   	OWF_Key[32,16]:=227126216;
   	OWF_Key[33,13]:=74826149;
   	OWF_Key[33,14]:=1639015971;
   	OWF_Key[33,15]:=305196101;
   	OWF_Key[33,16]:=716882039;
   	OWF_Key[34,13]:=380880877;
   	OWF_Key[34,14]:=11839263;
   	OWF_Key[34,15]:=1373141717;
   	OWF_Key[34,16]:=532627490;
   	OWF_Key[35,13]:=93438529;
   	OWF_Key[35,14]:=35115978;
   	OWF_Key[35,15]:=1081533615;
   	OWF_Key[35,16]:=1111729827;
   	OWF_Key[36,13]:=380331581;
   	OWF_Key[36,14]:=1532456188;
   	OWF_Key[36,15]:=1939052724;
   	OWF_Key[36,16]:=1794611672;
   	OWF_Key[37,13]:=1819289397;
   	OWF_Key[37,14]:=1027002065;
   	OWF_Key[37,15]:=1244500467;
   	OWF_Key[37,16]:=936638688;
   	OWF_Key[38,13]:=1479190277;
   	OWF_Key[38,14]:=519596430;
   	OWF_Key[38,15]:=1911107362;
   	OWF_Key[38,16]:=435044551;
   	OWF_Key[39,13]:=917290529;
   	OWF_Key[39,14]:=1617052636;
   	OWF_Key[39,15]:=606522633;
   	OWF_Key[39,16]:=1781888676;
   	OWF_Key[40,13]:=1628193547;
   	OWF_Key[40,14]:=89927245;
   	OWF_Key[40,15]:=820592385;
   	OWF_Key[40,16]:=524162027;
   	OWF_Key[41,13]:=699504604;
   	OWF_Key[41,14]:=2016929121;
   	OWF_Key[41,15]:=1410565984;
   	OWF_Key[41,16]:=1344454938;
   	OWF_Key[42,13]:=346920590;
   	OWF_Key[42,14]:=546121623;
   	OWF_Key[42,15]:=1947269171;
   	OWF_Key[42,16]:=311947312;
   	OWF_Key[43,13]:=673700248;
   	OWF_Key[43,14]:=2041423853;
   	OWF_Key[43,15]:=875126022;
   	OWF_Key[43,16]:=1745165237;
   	OWF_Key[44,13]:=1753633549;
   	OWF_Key[44,14]:=1140321993;
   	OWF_Key[44,15]:=33633727;
   	OWF_Key[44,16]:=1343682688;
   	OWF_Key[45,13]:=299201156;
   	OWF_Key[45,14]:=293335340;
   	OWF_Key[45,15]:=666355512;
   	OWF_Key[45,16]:=1885349377;
   	OWF_Key[46,13]:=1439159427;
   	OWF_Key[46,14]:=628092582;
   	OWF_Key[46,15]:=1364839979;
   	OWF_Key[46,16]:=1866912;
   	OWF_Key[47,13]:=856720789;
   	OWF_Key[47,14]:=930916762;
   	OWF_Key[47,15]:=2123174806;
   	OWF_Key[47,16]:=1671058401;
   	OWF_Key[48,13]:=230854938;
   	OWF_Key[48,14]:=878476914;
   	OWF_Key[48,15]:=1158749479;
   	OWF_Key[48,16]:=1143227675;
   	OWF_Key[49,13]:=2073892953;
   	OWF_Key[49,14]:=1273666786;
   	OWF_Key[49,15]:=2144362013;
   	OWF_Key[49,16]:=1099736956;
   	OWF_Key[50,13]:=874888610;
   	OWF_Key[50,14]:=1873711650;
   	OWF_Key[50,15]:=1719753255;
   	OWF_Key[50,16]:=1680711035;
   	OWF_Key[51,13]:=1361816747;
   	OWF_Key[51,14]:=1994614458;
   	OWF_Key[51,15]:=1199333913;
   	OWF_Key[51,16]:=1830471925;
   	OWF_Key[52,13]:=1995713668;
   	OWF_Key[52,14]:=919849947;
   	OWF_Key[52,15]:=767203999;
   	OWF_Key[52,16]:=1950347560;
   	OWF_Key[53,13]:=1787066567;
   	OWF_Key[53,14]:=1641494518;
   	OWF_Key[53,15]:=2137169354;
   	OWF_Key[53,16]:=1052747155;
   	OWF_Key[54,13]:=2054621143;
   	OWF_Key[54,14]:=1974715107;
   	OWF_Key[54,15]:=2111338725;
   	OWF_Key[54,16]:=1642760447;
   	OWF_Key[55,13]:=315851187;
   	OWF_Key[55,14]:=1955885849;
   	OWF_Key[55,15]:=2037754524;
   	OWF_Key[55,16]:=1309783764;
   	OWF_Key[56,13]:=629952185;
   	OWF_Key[56,14]:=210914935;
   	OWF_Key[56,15]:=1623244036;
   	OWF_Key[56,16]:=1765475415;
   	OWF_Key[57,13]:=857435203;
   	OWF_Key[57,14]:=206048520;
   	OWF_Key[57,15]:=369910258;
   	OWF_Key[57,16]:=1843731464;
   	OWF_Key[58,13]:=324501666;
   	OWF_Key[58,14]:=1733381472;
   	OWF_Key[58,15]:=1847843539;
   	OWF_Key[58,16]:=1608870174;
   	OWF_Key[59,13]:=1465774380;
   	OWF_Key[59,14]:=1286619525;
   	OWF_Key[59,15]:=573519412;
   	OWF_Key[59,16]:=1150347743;
   	OWF_Key[60,13]:=2015895654;
   	OWF_Key[60,14]:=201882130;
   	OWF_Key[60,15]:=1496789631;
   	OWF_Key[60,16]:=753620274;
   	OWF_Key[61,13]:=258623275;
   	OWF_Key[61,14]:=542640591;
   	OWF_Key[61,15]:=1506681182;
   	OWF_Key[61,16]:=1854703257;
   	OWF_Key[62,13]:=1141501595;
   	OWF_Key[62,14]:=1968246431;
   	OWF_Key[62,15]:=1731135653;
   	OWF_Key[62,16]:=2019442968;
   	OWF_Key[63,13]:=1282787873;
   	OWF_Key[63,14]:=579188533;
   	OWF_Key[63,15]:=1379806521;
   	OWF_Key[63,16]:=1195986330;
   	OWF_Key[64,13]:=1760745701;
   	OWF_Key[64,14]:=796682114;
   	OWF_Key[64,15]:=503806046;
   	OWF_Key[64,16]:=1014065369;
   	OWF_Key[65,13]:=744789352;
   	OWF_Key[65,14]:=1669355124;
   	OWF_Key[65,15]:=1249003689;
   	OWF_Key[65,16]:=446383216;
   	OWF_Key[66,13]:=1359397698;
   	OWF_Key[66,14]:=157427355;
   	OWF_Key[66,15]:=488697501;
   	OWF_Key[66,16]:=1040142022;
   	OWF_Key[67,13]:=881757290;
   	OWF_Key[67,14]:=965262803;
   	OWF_Key[67,15]:=1915722473;
   	OWF_Key[67,16]:=656835267;
   	OWF_Key[68,13]:=933499237;
   	OWF_Key[68,14]:=1187531747;
   	OWF_Key[68,15]:=197012920;
   	OWF_Key[68,16]:=274156957;
   	OWF_Key[69,13]:=1435849115;
   	OWF_Key[69,14]:=207728093;
   	OWF_Key[69,15]:=1550339381;
   	OWF_Key[69,16]:=924520084;
   	OWF_Key[70,13]:=1792435968;
   	OWF_Key[70,14]:=290098793;
   	OWF_Key[70,15]:=823633063;
   	OWF_Key[70,16]:=905749060;
   	OWF_Key[71,13]:=1550939045;
   	OWF_Key[71,14]:=2047053549;
   	OWF_Key[71,15]:=613147771;
   	OWF_Key[71,16]:=1592945744;
   	OWF_Key[72,13]:=1671761274;
   	OWF_Key[72,14]:=1866470197;
   	OWF_Key[72,15]:=1595615064;
   	OWF_Key[72,16]:=1624872080;
   	OWF_Key[73,13]:=1330706500;
   	OWF_Key[73,14]:=995552984;
   	OWF_Key[73,15]:=1155990823;
   	OWF_Key[73,16]:=166888145;
   	OWF_Key[74,13]:=935434492;
   	OWF_Key[74,14]:=1004579779;
   	OWF_Key[74,15]:=441645409;
   	OWF_Key[74,16]:=1173860650;
   	OWF_Key[75,13]:=124465085;
   	OWF_Key[75,14]:=1848317617;
   	OWF_Key[75,15]:=774434070;
   	OWF_Key[75,16]:=1822370621;
   	OWF_Key[76,13]:=1955710974;
   	OWF_Key[76,14]:=963579763;
   	OWF_Key[76,15]:=1302080192;
   	OWF_Key[76,16]:=1915358529;
   	OWF_Key[77,13]:=510947175;
   	OWF_Key[77,14]:=1670479738;
   	OWF_Key[77,15]:=658812905;
   	OWF_Key[77,16]:=6552539;
   	OWF_Key[78,13]:=958044673;
   	OWF_Key[78,14]:=381647451;
   	OWF_Key[78,15]:=510842397;
   	OWF_Key[78,16]:=916863139;
   	OWF_Key[79,13]:=127497795;
   	OWF_Key[79,14]:=806273643;
   	OWF_Key[79,15]:=1652287201;
   	OWF_Key[79,16]:=1761646512;
   	OWF_Key[80,13]:=1319108753;
   	OWF_Key[80,14]:=119208384;
   	OWF_Key[80,15]:=1872549858;
   	OWF_Key[80,16]:=1745731921;
   	OWF_Key[81,13]:=1435598528;
   	OWF_Key[81,14]:=571194510;
   	OWF_Key[81,15]:=191567415;
   	OWF_Key[81,16]:=217112706;
   	OWF_Key[82,13]:=1754599579;
   	OWF_Key[82,14]:=514829758;
   	OWF_Key[82,15]:=242412916;
   	OWF_Key[82,16]:=1451035335;
   	OWF_Key[83,13]:=1055894451;
   	OWF_Key[83,14]:=153938916;
   	OWF_Key[83,15]:=1360024240;
   	OWF_Key[83,16]:=398108754;
   	OWF_Key[84,13]:=1483905120;
   	OWF_Key[84,14]:=117806243;
   	OWF_Key[84,15]:=822813432;
   	OWF_Key[84,16]:=422563876;
   	OWF_Key[85,13]:=162587349;
   	OWF_Key[85,14]:=478421491;
   	OWF_Key[85,15]:=1015415493;
   	OWF_Key[85,16]:=1830070223;
   	OWF_Key[86,13]:=334994722;
   	OWF_Key[86,14]:=1913921160;
   	OWF_Key[86,15]:=1114283805;
   	OWF_Key[86,16]:=1127178650;
   	OWF_Key[87,13]:=1107170890;
   	OWF_Key[87,14]:=2012352564;
   	OWF_Key[87,15]:=57491098;
   	OWF_Key[87,16]:=1031931037;
   	OWF_Key[88,13]:=1840152318;
   	OWF_Key[88,14]:=1439707080;
   	OWF_Key[88,15]:=1204125942;
   	OWF_Key[88,16]:=460202532;
   	OWF_Key[89,13]:=357664832;
   	OWF_Key[89,14]:=651670053;
   	OWF_Key[89,15]:=949523032;
   	OWF_Key[89,16]:=30336271;
   	OWF_Key[90,13]:=1537181786;
   	OWF_Key[90,14]:=385729653;
   	OWF_Key[90,15]:=702817811;
   	OWF_Key[90,16]:=506086235;
   	OWF_Key[91,13]:=140712957;
   	OWF_Key[91,14]:=1989169662;
   	OWF_Key[91,15]:=1948213053;
   	OWF_Key[91,16]:=1066195582;
   	OWF_Key[92,13]:=1080088464;
   	OWF_Key[92,14]:=463170373;
   	OWF_Key[92,15]:=323347074;
   	OWF_Key[92,16]:=1133893629;
   	OWF_Key[93,13]:=908912253;
   	OWF_Key[93,14]:=551968720;
   	OWF_Key[93,15]:=1980909314;
   	OWF_Key[93,16]:=1712465128;
   	OWF_Key[94,13]:=1085647434;
   	OWF_Key[94,14]:=1044237653;
   	OWF_Key[94,15]:=1675868506;
   	OWF_Key[94,16]:=323851357;
   	OWF_Key[95,13]:=898355252;
   	OWF_Key[95,14]:=1501587080;
   	OWF_Key[95,15]:=1296328976;
   	OWF_Key[95,16]:=858795092;
   	OWF_Key[96,13]:=1480170052;
   	OWF_Key[96,14]:=1561016974;
   	OWF_Key[96,15]:=388658317;
   	OWF_Key[96,16]:=1336155871;
   	OWF_Key[97,13]:=347985099;
   	OWF_Key[97,14]:=1819162848;
   	OWF_Key[97,15]:=1472264812;
   	OWF_Key[97,16]:=638122137;
   	OWF_Key[98,13]:=1693384262;
   	OWF_Key[98,14]:=287561249;
   	OWF_Key[98,15]:=248517399;
   	OWF_Key[98,16]:=2033544562;
   	OWF_Key[99,13]:=440390558;
   	OWF_Key[99,14]:=1349263930;
   	OWF_Key[99,15]:=1752934582;
   	OWF_Key[99,16]:=1828420687;
   	OWF_Key[100,13]:=1779162509;
   	OWF_Key[100,14]:=147277535;
   	OWF_Key[100,15]:=1591203745;
   	OWF_Key[100,16]:=1387986523;
   	OWF_Key[101,13]:=893571876;
   	OWF_Key[101,14]:=1470481068;
   	OWF_Key[101,15]:=539793699;
   	OWF_Key[101,16]:=37186580;
   	OWF_Key[102,13]:=1710752197;
   	OWF_Key[102,14]:=1484165743;
   	OWF_Key[102,15]:=502723645;
   	OWF_Key[102,16]:=1327015877;
   	OWF_Key[103,13]:=812458487;
   	OWF_Key[103,14]:=1628876014;
   	OWF_Key[103,15]:=1328316236;
   	OWF_Key[103,16]:=2054343353;
   	OWF_Key[104,13]:=1919425969;
   	OWF_Key[104,14]:=896029992;
   	OWF_Key[104,15]:=1110917444;
   	OWF_Key[104,16]:=425290322;
   	OWF_Key[105,13]:=1924264538;
   	OWF_Key[105,14]:=1216674049;
   	OWF_Key[105,15]:=1533302189;
   	OWF_Key[105,16]:=2115098790;
   	OWF_Key[106,13]:=444126867;
   	OWF_Key[106,14]:=1038812109;
   	OWF_Key[106,15]:=1620113783;
   	OWF_Key[106,16]:=1670203207;
   	OWF_Key[107,13]:=853022640;
   	OWF_Key[107,14]:=1446113967;
   	OWF_Key[107,15]:=331193698;
   	OWF_Key[107,16]:=36897127;
   	OWF_Key[108,13]:=1772607745;
   	OWF_Key[108,14]:=278613042;
   	OWF_Key[108,15]:=1641923280;
   	OWF_Key[108,16]:=901128481;
   	OWF_Key[109,13]:=462107376;
   	OWF_Key[109,14]:=1753942874;
   	OWF_Key[109,15]:=1420322543;
   	OWF_Key[109,16]:=1585835244;
   	OWF_Key[110,13]:=1025292899;
   	OWF_Key[110,14]:=377139452;
   	OWF_Key[110,15]:=960310545;
   	OWF_Key[110,16]:=1455759124;
   	OWF_Key[111,13]:=978224434;
   	OWF_Key[111,14]:=1769099284;
   	OWF_Key[111,15]:=1469343786;
   	OWF_Key[111,16]:=1894157702;
   	OWF_Key[112,13]:=1579369767;
   	OWF_Key[112,14]:=1221710590;
   	OWF_Key[112,15]:=27970548;
   	OWF_Key[112,16]:=475176021;
   	OWF_Key[113,13]:=1406741878;
   	OWF_Key[113,14]:=1391221516;
   	OWF_Key[113,15]:=973931164;
   	OWF_Key[113,16]:=935798566;
   	OWF_Key[114,13]:=1016826153;
   	OWF_Key[114,14]:=395417869;
   	OWF_Key[114,15]:=139427492;
   	OWF_Key[114,16]:=380613091;
   	OWF_Key[115,13]:=1199001387;
   	OWF_Key[115,14]:=1643051957;
   	OWF_Key[115,15]:=867375944;
   	OWF_Key[115,16]:=1768598715;
   	OWF_Key[116,13]:=1371985039;
   	OWF_Key[116,14]:=239918248;
   	OWF_Key[116,15]:=475467365;
   	OWF_Key[116,16]:=352629576;
   	OWF_Key[117,13]:=406649522;
   	OWF_Key[117,14]:=1022185637;
   	OWF_Key[117,15]:=924251933;
   	OWF_Key[117,16]:=58287288;
   	OWF_Key[118,13]:=1444359901;
   	OWF_Key[118,14]:=1004398136;
   	OWF_Key[118,15]:=305939276;
   	OWF_Key[118,16]:=13282582;
   	OWF_Key[119,13]:=1753624650;
   	OWF_Key[119,14]:=395513408;
   	OWF_Key[119,15]:=1423144984;
   	OWF_Key[119,16]:=1539743838;
   	OWF_Key[120,13]:=442395067;
   	OWF_Key[120,14]:=2018925503;
   	OWF_Key[120,15]:=953917663;
   	OWF_Key[120,16]:=1688609331;
   	OWF_Key[121,13]:=787971890;
   	OWF_Key[121,14]:=1620287384;
   	OWF_Key[121,15]:=256968225;
   	OWF_Key[121,16]:=1301956638;
   	OWF_Key[122,13]:=990668381;
   	OWF_Key[122,14]:=2018680738;
   	OWF_Key[122,15]:=915563951;
   	OWF_Key[122,16]:=1304501418;
   	OWF_Key[123,13]:=845352878;
   	OWF_Key[123,14]:=1326819379;
   	OWF_Key[123,15]:=973867524;
   	OWF_Key[123,16]:=1330778393;
   	OWF_Key[124,13]:=1212459966;
   	OWF_Key[124,14]:=331345962;
   	OWF_Key[124,15]:=1503496153;
   	OWF_Key[124,16]:=1881291653;
   	OWF_Key[125,13]:=275083085;
   	OWF_Key[125,14]:=1241962392;
   	OWF_Key[125,15]:=1663659714;
   	OWF_Key[125,16]:=359811177;
   	OWF_Key[126,13]:=469249223;
   	OWF_Key[126,14]:=862227537;
   	OWF_Key[126,15]:=1043658105;
   	OWF_Key[126,16]:=1730970707;
   	OWF_Key[127,13]:=1168087958;
   	OWF_Key[127,14]:=282353341;
   	OWF_Key[127,15]:=343861148;
   	OWF_Key[127,16]:=2052225671;
   	OWF_Key[128,13]:=1557870208;
   	OWF_Key[128,14]:=1209923749;
   	OWF_Key[128,15]:=1776967874;
   	OWF_Key[128,16]:=288485818;
   	OWF_Key[129,13]:=74300695;
   	OWF_Key[129,14]:=968535377;
   	OWF_Key[129,15]:=851571720;
   	OWF_Key[129,16]:=2094292864;
   	OWF_Key[130,13]:=102777636;
   	OWF_Key[130,14]:=410444836;
   	OWF_Key[130,15]:=1304169589;
   	OWF_Key[130,16]:=1061853872;
   	OWF_Key[131,13]:=935817478;
   	OWF_Key[131,14]:=1893612138;
   	OWF_Key[131,15]:=462395237;
   	OWF_Key[131,16]:=681940591;
   	OWF_Key[132,13]:=381652625;
   	OWF_Key[132,14]:=201502794;
   	OWF_Key[132,15]:=1754047887;
   	OWF_Key[132,16]:=311395707;
   	OWF_Key[133,13]:=346211181;
   	OWF_Key[133,14]:=2071318594;
   	OWF_Key[133,15]:=1513459740;
   	OWF_Key[133,16]:=1115232146;
   	OWF_Key[134,13]:=1598695163;
   	OWF_Key[134,14]:=1466344949;
   	OWF_Key[134,15]:=762229445;
   	OWF_Key[134,16]:=672484557;
   	OWF_Key[135,13]:=1650533870;
   	OWF_Key[135,14]:=746136511;
   	OWF_Key[135,15]:=1403884082;
   	OWF_Key[135,16]:=1128504661;
   	OWF_Key[136,13]:=1193152325;
   	OWF_Key[136,14]:=1642319657;
   	OWF_Key[136,15]:=764561960;
   	OWF_Key[136,16]:=1782348027;
   	OWF_Key[137,13]:=481612577;
   	OWF_Key[137,14]:=1117357605;
   	OWF_Key[137,15]:=1226367764;
   	OWF_Key[137,16]:=486415909;
   	OWF_Key[138,13]:=712276525;
   	OWF_Key[138,14]:=1231818236;
   	OWF_Key[138,15]:=889849699;
   	OWF_Key[138,16]:=1322456834;
   	OWF_Key[139,13]:=1658882780;
   	OWF_Key[139,14]:=299855880;
   	OWF_Key[139,15]:=457182275;
   	OWF_Key[139,16]:=375856677;
   	OWF_Key[140,13]:=1427201989;
   	OWF_Key[140,14]:=1842532478;
   	OWF_Key[140,15]:=2020223672;
   	OWF_Key[140,16]:=95163959;
   	OWF_Key[141,13]:=1076016553;
   	OWF_Key[141,14]:=1900141535;
   	OWF_Key[141,15]:=1257026434;
   	OWF_Key[141,16]:=909049460;
   	OWF_Key[142,13]:=372483116;
   	OWF_Key[142,14]:=152435569;
   	OWF_Key[142,15]:=1367585177;
   	OWF_Key[142,16]:=180714971;
   	OWF_Key[143,13]:=492180917;
   	OWF_Key[143,14]:=811497737;
   	OWF_Key[143,15]:=182411329;
   	OWF_Key[143,16]:=1448390505;
   	OWF_Key[144,13]:=1474316502;
   	OWF_Key[144,14]:=962265029;
   	OWF_Key[144,15]:=2143233034;
   	OWF_Key[144,16]:=86163621;
   	OWF_Key[145,13]:=22318259;
   	OWF_Key[145,14]:=464103670;
   	OWF_Key[145,15]:=9486028;
   	OWF_Key[145,16]:=165100234;
   	OWF_Key[146,13]:=1738036540;
   	OWF_Key[146,14]:=957495089;
   	OWF_Key[146,15]:=1871584640;
   	OWF_Key[146,16]:=88784541;
   	OWF_Key[147,13]:=326829794;
   	OWF_Key[147,14]:=1163466676;
   	OWF_Key[147,15]:=1555104822;
   	OWF_Key[147,16]:=2103407692;
   	OWF_Key[148,13]:=1529543674;
   	OWF_Key[148,14]:=71476052;
   	OWF_Key[148,15]:=1157626873;
   	OWF_Key[148,16]:=1806721818;
   	OWF_Key[149,13]:=1849787839;
   	OWF_Key[149,14]:=931886575;
   	OWF_Key[149,15]:=657127511;
   	OWF_Key[149,16]:=1271697867;
   	OWF_Key[150,13]:=1381878125;
   	OWF_Key[150,14]:=1019077359;
   	OWF_Key[150,15]:=1860188757;
   	OWF_Key[150,16]:=1322712000;
   	OWF_Key[151,13]:=648949296;
   	OWF_Key[151,14]:=99719;
   	OWF_Key[151,15]:=1175680819;
   	OWF_Key[151,16]:=1497980896;
   	OWF_Key[152,13]:=1625442764;
   	OWF_Key[152,14]:=277771665;
   	OWF_Key[152,15]:=939669588;
   	OWF_Key[152,16]:=1601021974;
   	OWF_Key[153,13]:=899912740;
   	OWF_Key[153,14]:=251847340;
   	OWF_Key[153,15]:=549386803;
   	OWF_Key[153,16]:=800804065;
   	OWF_Key[154,13]:=1113652973;
   	OWF_Key[154,14]:=47019578;
   	OWF_Key[154,15]:=1748787020;
   	OWF_Key[154,16]:=1741961176;
   	OWF_Key[155,13]:=16858922;
   	OWF_Key[155,14]:=993261889;
   	OWF_Key[155,15]:=391546459;
   	OWF_Key[155,16]:=1613990827;
   	OWF_Key[156,13]:=359980847;
   	OWF_Key[156,14]:=17310265;
   	OWF_Key[156,15]:=992777913;
   	OWF_Key[156,16]:=1166263769;
   	OWF_Key[157,13]:=1948582787;
   	OWF_Key[157,14]:=281935467;
   	OWF_Key[157,15]:=1445300746;
   	OWF_Key[157,16]:=1211611796;
   	OWF_Key[158,13]:=178475878;
   	OWF_Key[158,14]:=202525481;
   	OWF_Key[158,15]:=131006593;
   	OWF_Key[158,16]:=1956785807;
   	OWF_Key[159,13]:=1801698601;
   	OWF_Key[159,14]:=726011192;
   	OWF_Key[159,15]:=1429967167;
   	OWF_Key[159,16]:=120231144;
   	OWF_Key[160,13]:=1755934677;
   	OWF_Key[160,14]:=931127830;
   	OWF_Key[160,15]:=1573768517;
   	OWF_Key[160,16]:=194947820;
   	OWF_Key[161,13]:=340873654;
   	OWF_Key[161,14]:=859703477;
   	OWF_Key[161,15]:=714867666;
   	OWF_Key[161,16]:=1308970684;
   	OWF_Key[162,13]:=2033262093;
   	OWF_Key[162,14]:=135322483;
   	OWF_Key[162,15]:=181185071;
   	OWF_Key[162,16]:=1019448048;
   	OWF_Key[163,13]:=351815141;
   	OWF_Key[163,14]:=1349943554;
   	OWF_Key[163,15]:=1519426241;
   	OWF_Key[163,16]:=1730005141;
   	OWF_Key[164,13]:=895515385;
   	OWF_Key[164,14]:=759942475;
   	OWF_Key[164,15]:=1274974076;
   	OWF_Key[164,16]:=1778058459;
   	OWF_Key[165,13]:=1534002997;
   	OWF_Key[165,14]:=342683598;
   	OWF_Key[165,15]:=1325035008;
   	OWF_Key[165,16]:=541951738;
   	OWF_Key[166,13]:=1126159679;
   	OWF_Key[166,14]:=1135178360;
   	OWF_Key[166,15]:=171444871;
   	OWF_Key[166,16]:=1500118001;
   	OWF_Key[167,13]:=1319550750;
   	OWF_Key[167,14]:=1523155912;
   	OWF_Key[167,15]:=1894915506;
   	OWF_Key[167,16]:=46108147;
   	OWF_Key[168,13]:=891586055;
   	OWF_Key[168,14]:=1614220493;
   	OWF_Key[168,15]:=948985067;
   	OWF_Key[168,16]:=1008303949;
   	OWF_Key[169,13]:=714425471;
   	OWF_Key[169,14]:=404425965;
   	OWF_Key[169,15]:=1214720770;
   	OWF_Key[169,16]:=661094727;
   	OWF_Key[170,13]:=1417632945;
   	OWF_Key[170,14]:=1553623603;
   	OWF_Key[170,15]:=1142877093;
   	OWF_Key[170,16]:=1852102698;
   	OWF_Key[171,13]:=1325459671;
   	OWF_Key[171,14]:=1213428668;
   	OWF_Key[171,15]:=791381338;
   	OWF_Key[171,16]:=1093670539;
   	OWF_Key[172,13]:=67122307;
   	OWF_Key[172,14]:=722754093;
   	OWF_Key[172,15]:=1643848423;
   	OWF_Key[172,16]:=830718530;
   	OWF_Key[173,13]:=984850756;
   	OWF_Key[173,14]:=1149842119;
   	OWF_Key[173,15]:=171832428;
   	OWF_Key[173,16]:=2085848996;
   	OWF_Key[174,13]:=1995806419;
   	OWF_Key[174,14]:=811214497;
   	OWF_Key[174,15]:=1118289432;
   	OWF_Key[174,16]:=726787119;
   	OWF_Key[175,13]:=372222373;
   	OWF_Key[175,14]:=946921363;
   	OWF_Key[175,15]:=1763664559;
   	OWF_Key[175,16]:=1522951892;
   	OWF_Key[176,13]:=753425289;
   	OWF_Key[176,14]:=1971291402;
   	OWF_Key[176,15]:=1757383876;
   	OWF_Key[176,16]:=554600741;
   	OWF_Key[177,13]:=2116933958;
   	OWF_Key[177,14]:=684392856;
   	OWF_Key[177,15]:=1940251711;
   	OWF_Key[177,16]:=48359718;
   	OWF_Key[178,13]:=2028009177;
   	OWF_Key[178,14]:=48868902;
   	OWF_Key[178,15]:=89820102;
   	OWF_Key[178,16]:=1140097925;
   	OWF_Key[179,13]:=1985450806;
   	OWF_Key[179,14]:=1466515194;
   	OWF_Key[179,15]:=1981559753;
   	OWF_Key[179,16]:=465352035;
   	OWF_Key[180,13]:=1999606185;
   	OWF_Key[180,14]:=824765067;
   	OWF_Key[180,15]:=389379872;
   	OWF_Key[180,16]:=334105230;
   	OWF_Key[181,13]:=1123156879;
   	OWF_Key[181,14]:=1288903172;
   	OWF_Key[181,15]:=588243473;
   	OWF_Key[181,16]:=377190400;
   	OWF_Key[182,13]:=331455980;
   	OWF_Key[182,14]:=757004017;
   	OWF_Key[182,15]:=1679453652;
   	OWF_Key[182,16]:=953675030;
   	OWF_Key[183,13]:=319703761;
   	OWF_Key[183,14]:=686929024;
   	OWF_Key[183,15]:=1771394380;
   	OWF_Key[183,16]:=1146391459;
   	OWF_Key[184,13]:=64113331;
   	OWF_Key[184,14]:=1843233077;
   	OWF_Key[184,15]:=1054710883;
   	OWF_Key[184,16]:=16307061;
   	OWF_Key[185,13]:=577790918;
   	OWF_Key[185,14]:=769951951;
   	OWF_Key[185,15]:=36875238;
   	OWF_Key[185,16]:=969551747;
   	OWF_Key[186,13]:=1949099229;
   	OWF_Key[186,14]:=16345749;
   	OWF_Key[186,15]:=1812777874;
   	OWF_Key[186,16]:=1770825016;
   	OWF_Key[187,13]:=360969632;
   	OWF_Key[187,14]:=1677985071;
   	OWF_Key[187,15]:=1100521128;
   	OWF_Key[187,16]:=1658272940;
   	OWF_Key[188,13]:=1778139981;
   	OWF_Key[188,14]:=1202793776;
   	OWF_Key[188,15]:=17874512;
   	OWF_Key[188,16]:=2077025197;
   	OWF_Key[189,13]:=1605074632;
   	OWF_Key[189,14]:=735118058;
   	OWF_Key[189,15]:=2120994248;
   	OWF_Key[189,16]:=1327201891;
   	OWF_Key[190,13]:=2070065568;
   	OWF_Key[190,14]:=1393044672;
   	OWF_Key[190,15]:=976654796;
   	OWF_Key[190,16]:=1710671530;
   	OWF_Key[191,13]:=38568234;
   	OWF_Key[191,14]:=451698160;
   	OWF_Key[191,15]:=1261954091;
   	OWF_Key[191,16]:=249271037;
   	OWF_Key[192,13]:=1638949335;
   	OWF_Key[192,14]:=8243760;
   	OWF_Key[192,15]:=241234447;
   	OWF_Key[192,16]:=1227077516;
   	OWF_Key[193,13]:=989587635;
   	OWF_Key[193,14]:=1819989847;
   	OWF_Key[193,15]:=1332579048;
   	OWF_Key[193,16]:=53755968;
   	OWF_Key[194,13]:=100673663;
   	OWF_Key[194,14]:=1469329794;
   	OWF_Key[194,15]:=1436971146;
   	OWF_Key[194,16]:=929174323;
   	OWF_Key[195,13]:=577996306;
   	OWF_Key[195,14]:=1745684579;
   	OWF_Key[195,15]:=1996965839;
   	OWF_Key[195,16]:=1403732815;
   	OWF_Key[196,13]:=814419608;
   	OWF_Key[196,14]:=2103643129;
   	OWF_Key[196,15]:=335105042;
   	OWF_Key[196,16]:=565961710;
   	OWF_Key[197,13]:=202009593;
   	OWF_Key[197,14]:=930351125;
   	OWF_Key[197,15]:=1526609745;
   	OWF_Key[197,16]:=235969148;
   	OWF_Key[198,13]:=1626921131;
   	OWF_Key[198,14]:=161315506;
   	OWF_Key[198,15]:=767020089;
   	OWF_Key[198,16]:=624440912;
   	OWF_Key[199,13]:=684936633;
   	OWF_Key[199,14]:=1742723201;
   	OWF_Key[199,15]:=515114070;
   	OWF_Key[199,16]:=162561603;
   	OWF_Key[200,13]:=1845652691;
   	OWF_Key[200,14]:=1950369016;
   	OWF_Key[200,15]:=571396495;
   	OWF_Key[200,16]:=1488194196;
   	OWF_Key[201,13]:=1043958765;
   	OWF_Key[201,14]:=1442574514;
   	OWF_Key[201,15]:=298914684;
   	OWF_Key[201,16]:=486285287;
   	OWF_Key[202,13]:=1582775329;
   	OWF_Key[202,14]:=838793472;
   	OWF_Key[202,15]:=418382333;
   	OWF_Key[202,16]:=10776897;
   	OWF_Key[203,13]:=356986201;
   	OWF_Key[203,14]:=1108865874;
   	OWF_Key[203,15]:=1219664864;
   	OWF_Key[203,16]:=333594191;
   	OWF_Key[204,13]:=1541947490;
   	OWF_Key[204,14]:=1287551736;
   	OWF_Key[204,15]:=2059108066;
   	OWF_Key[204,16]:=1345707128;
   	OWF_Key[205,13]:=471367747;
   	OWF_Key[205,14]:=1525775149;
   	OWF_Key[205,15]:=1316108369;
   	OWF_Key[205,16]:=204019700;
   	OWF_Key[206,13]:=1473740948;
   	OWF_Key[206,14]:=286079449;
   	OWF_Key[206,15]:=1267750516;
   	OWF_Key[206,16]:=1937545157;
   	OWF_Key[207,13]:=2126324793;
   	OWF_Key[207,14]:=1789210342;
   	OWF_Key[207,15]:=501529746;
   	OWF_Key[207,16]:=2059785685;
   	OWF_Key[208,13]:=1274331883;
   	OWF_Key[208,14]:=968436149;
   	OWF_Key[208,15]:=1212562234;
   	OWF_Key[208,16]:=1455603155;
   	OWF_Key[209,13]:=92139053;
   	OWF_Key[209,14]:=992103779;
   	OWF_Key[209,15]:=1748163220;
   	OWF_Key[209,16]:=1233220835;
   	OWF_Key[210,13]:=259332684;
   	OWF_Key[210,14]:=2097850167;
   	OWF_Key[210,15]:=1049341383;
   	OWF_Key[210,16]:=714331988;
   	OWF_Key[211,13]:=1943218259;
   	OWF_Key[211,14]:=783610855;
   	OWF_Key[211,15]:=1161953504;
   	OWF_Key[211,16]:=1696436050;
   	OWF_Key[212,13]:=153726579;
   	OWF_Key[212,14]:=1993949032;
   	OWF_Key[212,15]:=281746886;
   	OWF_Key[212,16]:=2143629952;
   	OWF_Key[213,13]:=605671393;
   	OWF_Key[213,14]:=1472561361;
   	OWF_Key[213,15]:=1039695812;
   	OWF_Key[213,16]:=1849168053;
   	OWF_Key[214,13]:=1769778486;
   	OWF_Key[214,14]:=45741824;
   	OWF_Key[214,15]:=87024642;
   	OWF_Key[214,16]:=327652964;
   	OWF_Key[215,13]:=1490125572;
   	OWF_Key[215,14]:=1994649884;
   	OWF_Key[215,15]:=1234571844;
   	OWF_Key[215,16]:=920030323;
   	OWF_Key[216,13]:=2133174690;
   	OWF_Key[216,14]:=95558060;
   	OWF_Key[216,15]:=615326818;
   	OWF_Key[216,16]:=761728021;
   	OWF_Key[217,13]:=382282573;
   	OWF_Key[217,14]:=2017861784;
   	OWF_Key[217,15]:=1878700514;
   	OWF_Key[217,16]:=1515922417;
   	OWF_Key[218,13]:=1408298373;
   	OWF_Key[218,14]:=2039732974;
   	OWF_Key[218,15]:=1146678000;
   	OWF_Key[218,16]:=527275423;
   	OWF_Key[219,13]:=9291349;
   	OWF_Key[219,14]:=1702428079;
   	OWF_Key[219,15]:=340543343;
   	OWF_Key[219,16]:=1326649665;
   	OWF_Key[220,13]:=688341233;
   	OWF_Key[220,14]:=641189597;
   	OWF_Key[220,15]:=909299166;
   	OWF_Key[220,16]:=1752870415;
   	OWF_Key[221,13]:=1293014471;
   	OWF_Key[221,14]:=1168109613;
   	OWF_Key[221,15]:=1639198412;
   	OWF_Key[221,16]:=1211155230;
   	OWF_Key[222,13]:=1094302685;
   	OWF_Key[222,14]:=1748380807;
   	OWF_Key[222,15]:=740974356;
   	OWF_Key[222,16]:=981054882;
   	OWF_Key[223,13]:=1672948985;
   	OWF_Key[223,14]:=653486474;
   	OWF_Key[223,15]:=252491540;
   	OWF_Key[223,16]:=233857892;
   	OWF_Key[224,13]:=1488948359;
   	OWF_Key[224,14]:=855793400;
   	OWF_Key[224,15]:=299892487;
   	OWF_Key[224,16]:=955554724;
   	OWF_Key[225,13]:=1321934707;
   	OWF_Key[225,14]:=515714607;
   	OWF_Key[225,15]:=1346403512;
   	OWF_Key[225,16]:=540889864;
   	OWF_Key[226,13]:=760856919;
   	OWF_Key[226,14]:=452777885;
   	OWF_Key[226,15]:=152820366;
   	OWF_Key[226,16]:=158283786;
   	OWF_Key[227,13]:=1089442553;
   	OWF_Key[227,14]:=2136824552;
   	OWF_Key[227,15]:=492274941;
   	OWF_Key[227,16]:=1279116002;
   	OWF_Key[228,13]:=1639087779;
   	OWF_Key[228,14]:=1218708088;
   	OWF_Key[228,15]:=1350789742;
   	OWF_Key[228,16]:=266569552;
   	OWF_Key[229,13]:=63735330;
   	OWF_Key[229,14]:=1886757000;
   	OWF_Key[229,15]:=1923484766;
   	OWF_Key[229,16]:=1872440511;
   	OWF_Key[230,13]:=1943052252;
   	OWF_Key[230,14]:=1939759099;
   	OWF_Key[230,15]:=1108124166;
   	OWF_Key[230,16]:=1825389873;
   	OWF_Key[231,13]:=106697806;
   	OWF_Key[231,14]:=934330632;
   	OWF_Key[231,15]:=1226706106;
   	OWF_Key[231,16]:=1350717017;
   	OWF_Key[232,13]:=894995339;
   	OWF_Key[232,14]:=351973824;
   	OWF_Key[232,15]:=1915615287;
   	OWF_Key[232,16]:=1129455312;
   	OWF_Key[233,13]:=1606628665;
   	OWF_Key[233,14]:=792183115;
   	OWF_Key[233,15]:=655199967;
   	OWF_Key[233,16]:=466042394;
   	OWF_Key[234,13]:=265845209;
   	OWF_Key[234,14]:=1445558412;
   	OWF_Key[234,15]:=929515350;
   	OWF_Key[234,16]:=1736036285;
   	OWF_Key[235,13]:=1417713492;
   	OWF_Key[235,14]:=1710605342;
   	OWF_Key[235,15]:=153446933;
   	OWF_Key[235,16]:=200651284;
   	OWF_Key[236,13]:=1199064634;
   	OWF_Key[236,14]:=1304667317;
   	OWF_Key[236,15]:=1611340556;
   	OWF_Key[236,16]:=1688220347;
   	OWF_Key[237,13]:=1064686683;
   	OWF_Key[237,14]:=808058326;
   	OWF_Key[237,15]:=602176291;
   	OWF_Key[237,16]:=1592512372;
   	OWF_Key[238,13]:=188870782;
   	OWF_Key[238,14]:=699286542;
   	OWF_Key[238,15]:=740512834;
   	OWF_Key[238,16]:=805888291;
   	OWF_Key[239,13]:=2112249627;
   	OWF_Key[239,14]:=104687811;
   	OWF_Key[239,15]:=327040909;
   	OWF_Key[239,16]:=106310827;
   	OWF_Key[240,13]:=1922545948;
   	OWF_Key[240,14]:=1158736547;
   	OWF_Key[240,15]:=1646338950;
   	OWF_Key[240,16]:=302904535;
   	OWF_Key[241,13]:=1445166756;
   	OWF_Key[241,14]:=619904940;
   	OWF_Key[241,15]:=805963919;
   	OWF_Key[241,16]:=1775549581;
   	OWF_Key[242,13]:=461521008;
   	OWF_Key[242,14]:=1556197099;
   	OWF_Key[242,15]:=1292972172;
   	OWF_Key[242,16]:=1092790932;
   	OWF_Key[243,13]:=1366207430;
   	OWF_Key[243,14]:=1785310964;
   	OWF_Key[243,15]:=568468368;
   	OWF_Key[243,16]:=1252968121;
   	OWF_Key[244,13]:=973501638;
   	OWF_Key[244,14]:=859732749;
   	OWF_Key[244,15]:=1833062061;
   	OWF_Key[244,16]:=572987018;
   	OWF_Key[245,13]:=791865080;
   	OWF_Key[245,14]:=1765055225;
   	OWF_Key[245,15]:=310873594;
   	OWF_Key[245,16]:=589255605;
   	OWF_Key[246,13]:=1759833367;
   	OWF_Key[246,14]:=1618489300;
   	OWF_Key[246,15]:=830573894;
   	OWF_Key[246,16]:=1046861291;
   	OWF_Key[247,13]:=273538380;
   	OWF_Key[247,14]:=45619103;
   	OWF_Key[247,15]:=1158253128;
   	OWF_Key[247,16]:=142007761;
   	OWF_Key[248,13]:=307057508;
   	OWF_Key[248,14]:=1407424654;
   	OWF_Key[248,15]:=1570069593;
   	OWF_Key[248,16]:=832481957;
   	OWF_Key[249,13]:=962494443;
   	OWF_Key[249,14]:=1117874804;
   	OWF_Key[249,15]:=1823842561;
   	OWF_Key[249,16]:=1850442054;
   	OWF_Key[250,13]:=1442058163;
   	OWF_Key[250,14]:=1232560055;
   	OWF_Key[250,15]:=151821927;
   	OWF_Key[250,16]:=1056371398;
   	OWF_Key[251,13]:=332739772;
   	OWF_Key[251,14]:=2051033636;
   	OWF_Key[251,15]:=849642509;
   	OWF_Key[251,16]:=1992496557;
   	OWF_Key[252,13]:=1955024293;
   	OWF_Key[252,14]:=864654120;
   	OWF_Key[252,15]:=400202456;
   	OWF_Key[252,16]:=1469872697;
   	OWF_Key[253,13]:=1814679055;
   	OWF_Key[253,14]:=1018947711;
   	OWF_Key[253,15]:=414056628;
   	OWF_Key[253,16]:=1916175716;
   	OWF_Key[254,13]:=34988910;
   	OWF_Key[254,14]:=1068930085;
   	OWF_Key[254,15]:=1069419481;
   	OWF_Key[254,16]:=1329460403;
   	OWF_Key[255,13]:=629578987;
   	OWF_Key[255,14]:=1913112785;
   	OWF_Key[255,15]:=1118884227;
   	OWF_Key[255,16]:=660504630;
   	OWF_Key[256,13]:=1745889977;
   	OWF_Key[256,14]:=1744367642;
   	OWF_Key[256,15]:=1635265674;
   	OWF_Key[256,16]:=250591589;
   	OWF_Key[257,13]:=1359647390;
   	OWF_Key[257,14]:=335557629;
   	OWF_Key[257,15]:=272575744;
   	OWF_Key[257,16]:=782479111;
   	OWF_Key[258,13]:=1684017798;
   	OWF_Key[258,14]:=1849154465;
   	OWF_Key[258,15]:=131467400;
   	OWF_Key[258,16]:=244488627;
   	OWF_Key[259,13]:=41240583;
   	OWF_Key[259,14]:=963084835;
   	OWF_Key[259,15]:=844053562;
   	OWF_Key[259,16]:=1313394598;
   	OWF_Key[260,13]:=646795143;
   	OWF_Key[260,14]:=1614027852;
   	OWF_Key[260,15]:=2028202305;
   	OWF_Key[260,16]:=1145473513;
   	OWF_Key[261,13]:=16520506;
   	OWF_Key[261,14]:=1480547316;
   	OWF_Key[261,15]:=1576651890;
   	OWF_Key[261,16]:=326846098;
   	OWF_Key[262,13]:=274761447;
   	OWF_Key[262,14]:=981162513;
   	OWF_Key[262,15]:=960880365;
   	OWF_Key[262,16]:=535655077;
   	OWF_Key[263,13]:=815853165;
   	OWF_Key[263,14]:=965917766;
   	OWF_Key[263,15]:=1914171172;
   	OWF_Key[263,16]:=192053027;
   	OWF_Key[264,13]:=908824118;
   	OWF_Key[264,14]:=2075268001;
   	OWF_Key[264,15]:=314233580;
   	OWF_Key[264,16]:=1793819686;
   	OWF_Key[265,13]:=928633642;
   	OWF_Key[265,14]:=1394677407;
   	OWF_Key[265,15]:=381077257;
   	OWF_Key[265,16]:=1427933170;
   	OWF_Key[266,13]:=1325823149;
   	OWF_Key[266,14]:=326658029;
   	OWF_Key[266,15]:=1415638516;
   	OWF_Key[266,16]:=1370549208;
   	OWF_Key[267,13]:=91918653;
   	OWF_Key[267,14]:=1189442786;
   	OWF_Key[267,15]:=1488204864;
   	OWF_Key[267,16]:=739198522;
   	OWF_Key[268,13]:=1461502145;
   	OWF_Key[268,14]:=84921185;
   	OWF_Key[268,15]:=440014277;
   	OWF_Key[268,16]:=2099928856;
   	OWF_Key[269,13]:=1927983756;
   	OWF_Key[269,14]:=1119840967;
   	OWF_Key[269,15]:=388770855;
   	OWF_Key[269,16]:=1179250891;
   	OWF_Key[270,13]:=126605253;
   	OWF_Key[270,14]:=777231285;
   	OWF_Key[270,15]:=2005758675;
   	OWF_Key[270,16]:=1335960631;
   	OWF_Key[271,13]:=1845648579;
   	OWF_Key[271,14]:=380266852;
   	OWF_Key[271,15]:=248475413;
   	OWF_Key[271,16]:=331001610;
   	OWF_Key[272,13]:=605803683;
   	OWF_Key[272,14]:=607759287;
   	OWF_Key[272,15]:=665317173;
   	OWF_Key[272,16]:=1066666071;
   	OWF_Key[273,13]:=1398348673;
   	OWF_Key[273,14]:=848648801;
   	OWF_Key[273,15]:=867913242;
   	OWF_Key[273,16]:=138992559;
   	OWF_Key[274,13]:=610350804;
   	OWF_Key[274,14]:=523330815;
   	OWF_Key[274,15]:=1415166854;
   	OWF_Key[274,16]:=1770062347;
   	OWF_Key[275,13]:=835727048;
   	OWF_Key[275,14]:=35430845;
   	OWF_Key[275,15]:=596122974;
   	OWF_Key[275,16]:=684344241;
   	OWF_Key[276,13]:=78641305;
   	OWF_Key[276,14]:=788905719;
   	OWF_Key[276,15]:=880092642;
   	OWF_Key[276,16]:=1020585456;
   	OWF_Key[277,13]:=1110913439;
   	OWF_Key[277,14]:=1364792795;
   	OWF_Key[277,15]:=1384151855;
   	OWF_Key[277,16]:=1781215518;
   	OWF_Key[278,13]:=1664996503;
   	OWF_Key[278,14]:=1954790028;
   	OWF_Key[278,15]:=320064116;
   	OWF_Key[278,16]:=318277611;
   	OWF_Key[279,13]:=1474869755;
   	OWF_Key[279,14]:=1993904309;
   	OWF_Key[279,15]:=749636549;
   	OWF_Key[279,16]:=2065511657;
   	OWF_Key[280,13]:=903827560;
   	OWF_Key[280,14]:=1827376749;
   	OWF_Key[280,15]:=103307236;
   	OWF_Key[280,16]:=510364959;
   	OWF_Key[281,13]:=1734942199;
   	OWF_Key[281,14]:=442316326;
   	OWF_Key[281,15]:=1226640256;
   	OWF_Key[281,16]:=668862109;
   	OWF_Key[282,13]:=218310287;
   	OWF_Key[282,14]:=528444193;
   	OWF_Key[282,15]:=1586604669;
   	OWF_Key[282,16]:=63254231;
   	OWF_Key[283,13]:=689997306;
   	OWF_Key[283,14]:=1451778241;
   	OWF_Key[283,15]:=2105293635;
   	OWF_Key[283,16]:=1663094505;
   	OWF_Key[284,13]:=1377189714;
   	OWF_Key[284,14]:=1670984675;
   	OWF_Key[284,15]:=309287320;
   	OWF_Key[284,16]:=1604200948;
   	OWF_Key[285,13]:=709339406;
   	OWF_Key[285,14]:=1683608969;
   	OWF_Key[285,15]:=109866542;
   	OWF_Key[285,16]:=480182101;
   	OWF_Key[286,13]:=1653006727;
   	OWF_Key[286,14]:=1931713950;
   	OWF_Key[286,15]:=221605941;
   	OWF_Key[286,16]:=859421666;
   	OWF_Key[287,13]:=1624256019;
   	OWF_Key[287,14]:=1737854557;
   	OWF_Key[287,15]:=199703631;
   	OWF_Key[287,16]:=428542639;
   	OWF_Key[288,13]:=1395232127;
   	OWF_Key[288,14]:=441805761;
   	OWF_Key[288,15]:=1127303696;
   	OWF_Key[288,16]:=544157041;
   	OWF_Key[289,13]:=1812633173;
   	OWF_Key[289,14]:=703745186;
